(* Logix 5000 project; controller FV vendor 1 type 14 code 217 rev 31.11; software revision 31.00; part 62 of 63 *)
(* tags used below, declared in another part *)
   CWD : CHECKWORD_FLAGS;
   YP_AV1 : PlantItem;   // AV1
   YP_AV2 : PlantItem;   // AV2
   YP_AV3 : PlantItem;   // AV3
   YP_AV4 : PlantItem;   // AV4
   YP_AV5 : PlantItem;   // AV5
   YP_AV6 : PlantItem;   // AV6
   YP_AV7 : PlantItem;   // AV7
   YP_AV8 : PlantItem;   // AV8
   YP_B103 : INT[15];   // Original N File From SLC, No Description Available
   YP_B3 : INT[7];   // BINARY
   YP_B30 : INT[37];   // Original N File From SLC, No Description Available
   YP_B92 : INT[105];   // Original N File From SLC, No Description Available
   YP_BLUNG_OV : PlantItem;   // BLUNG_OV
   YP_C5 : COUNTER[15];
   YP_COMMS_FROM_MVFVCIP : MESSAGE;
   YP_CONV_STOP : PlantItem;   // CONV_STOP
   YP_INP1 : PlantItem;   // INP1
   YP_INP10 : PlantItem;   // INP10
   YP_INP11 : PlantItem;   // INP11
   YP_INP2 : PlantItem;   // INP2
   YP_INP3 : PlantItem;   // INP3
   YP_INP4 : PlantItem;   // INP4
   YP_INP5 : PlantItem;   // INP5
   YP_INP6 : PlantItem;   // INP6
   YP_INP7 : PlantItem;   // INP7
   YP_INP8 : PlantItem;   // INP8
   YP_INP9 : PlantItem;   // INP9
   YP_N14 : INT[135];   // Original N File From SLC, No Description Available
   YP_N40 : INT[9];   // Original N File From SLC, No Description Available
   YP_N55 : INT[244];   // Original N File From SLC, No Description Available
   YP_OUT1 : PlantItem;   // OUT1
   YP_OUT2 : PlantItem;   // OUT2
   YP_OUT3 : PlantItem;   // OUT3
   YP_OUT4 : PlantItem;   // OUT4
   YP_OUT5 : PlantItem;   // OUT5
   YP_OUT6 : PlantItem;   // OUT6
   YP_OUT7 : PlantItem;   // OUT7
   YP_PILZ_OK : PlantItem;   // PILZ_OK
   YP_PRESS_CL : PlantItem;   // PRESS_CL
   YP_PRESS_OP : PlantItem;   // PRESS_OP
   YP_T21 : TIMER[30];
   YP_T4 : TIMER[16];   // TIMER
   YP_WD : PlantItem;   // WD
   YP_WD_RawOutput : ALIAS FOR RIO_Rack_3:3:O.Data.14;   // YP_WD
   YST_BL_PMP_ON : BOOL;   // Blunger Pump
(* YP_Common, continued *)

ROUTINE YP_Digital_Outputs   (* ladder *)
   0: [NEQ(YP_WD.DriveBits,0) OTE(YP_WD.CW.[CWD.AUTODRV]) ,XIC(S:FS) OTU(YP_WD.CW.[CWD.MANUAL]) ,[XIC(YP_WD.CW.[CWD.AUTODRV]) XIO(YP_WD.CW.[CWD.MANUAL]) ,XIC(YP_WD.CW.[CWD.MANDRV]) XIC(YP_WD.CW.[CWD.MANUAL]) ] OTE(YP_WD.CW.[CWD.OUTPUT]) ,XIC(YP_WD.CW.[CWD.OUTPUT]) OTE(YP_WD_RawOutput) ];
END_ROUTINE

ROUTINE YP_INPUTS_10   (* ladder *)
   0: XIC(YP_AV1.CW.[CWD.OPENFB])OTE(YP_B3[0].0);
   1: XIC(YP_AV2.CW.[CWD.OPENFB])OTE(YP_B3[0].2);
   2: XIC(YP_AV3.CW.[CWD.OPENFB])OTE(YP_B3[0].4);
   3: XIC(YP_AV4.CW.[CWD.OPENFB])OTE(YP_B3[0].6);
   4: XIC(YP_AV5.CW.[CWD.OPENFB])OTE(YP_B3[0].8);
   5: XIC(YP_AV6.CW.[CWD.OPENFB])OTE(YP_B3[0].10);
   6: XIC(YP_AV7.CW.[CWD.OPENFB])OTE(YP_B3[0].12);
   7: XIC(YP_AV8.CW.[CWD.OPENFB])OTE(YP_B3[0].14);
   8: XIC(YP_PILZ_OK.CW.[CWD.INPUTSTATUS])OTE(YP_B3[1].0);
   9: XIC(YP_BLUNG_OV.CW.[CWD.INPUTSTATUS])OTE(YP_B3[1].1);
   10: XIO(YP_INP1.CW.[CWD.INPUTSTATUS])OTE(YP_B3[1].2);
   11: XIC(YP_INP2.CW.[CWD.INPUTSTATUS])OTE(YP_B3[1].3);
   12: XIC(YP_INP3.CW.[CWD.INPUTSTATUS])OTE(YP_B3[1].4);
   13: XIC(YP_PRESS_CL.CW.[CWD.INPUTSTATUS])OTE(YP_B3[1].5);
   14: XIC(YP_PRESS_OP.CW.[CWD.INPUTSTATUS])OTE(YP_B3[1].6);
   15: XIC(YP_CONV_STOP.CW.[CWD.INPUTSTATUS])OTE(YP_B3[1].7);
   16: XIC(YP_INP4.CW.[CWD.INPUTSTATUS])OTE(YP_B3[1].8);
   17: XIC(YP_INP5.CW.[CWD.INPUTSTATUS])OTE(YP_B3[1].9);
   18: XIC(YP_INP6.CW.[CWD.INPUTSTATUS])OTE(YP_B3[1].10);
   19: XIC(YP_INP7.CW.[CWD.INPUTSTATUS])OTE(YP_B3[1].11);
   20: XIC(YP_INP8.CW.[CWD.INPUTSTATUS])OTE(YP_B3[1].12);
   21: XIC(YP_INP9.CW.[CWD.INPUTSTATUS])OTE(YP_B3[1].13);
   22: XIC(YP_INP10.CW.[CWD.INPUTSTATUS])OTE(YP_B3[1].14);
   23: XIC(YP_INP11.CW.[CWD.INPUTSTATUS])OTE(YP_B3[1].15);
END_ROUTINE

ROUTINE YP_LAD15_15   (* ladder *)
   0: XIO(YP_T4[3].DN)TON(YP_T4[3],?,?);
   1: XIO(YP_N40[0].0)XIO(YP_N40[0].1)XIO(YP_N40[0].2)XIO(YP_N40[0].3)XIO(YP_N40[0].4)XIO(YP_N40[0].5)XIO(YP_N40[0].6)XIO(YP_N40[0].7)XIO(YP_N40[0].8)[OTL(YP_N40[0].0) ,OTU(YP_N40[0].1) ,OTU(YP_N40[0].2) ,OTU(YP_N40[0].3) ,OTU(YP_N40[0].4) ,OTU(YP_N40[0].5) ,OTU(YP_N40[0].6) ,OTU(YP_N40[0].7) ,OTU(YP_N40[0].8) ];
   2: XIC(YP_N40[0].8)XIC(YP_B3[1].7)[OTU(YP_N40[0].8) ,OTL(YP_N40[0].0) ];
   3: XIC(YP_N40[0].0)XIC(YP_B3[1].0)XIC(YP_B3[1].5)EQU(YP_N55[0],0)[OTU(YP_N40[0].0) ,OTL(YP_N40[0].1) ];
   4: XIC(YP_N40[0].1)XIC(YP_B3[1].1)[OTU(YP_N40[0].1) ,OTL(YP_N40[0].2) ];
   5: XIC(YP_N40[0].2)TON(YP_T21[0],?,?);
   6: XIC(YP_N40[0].2)XIC(YP_T21[0].DN)[OTU(YP_N40[0].2) ,OTL(YP_N40[0].3) ];
   7: MOV(YP_N55[20],YP_C5[0].PRE);
   8: XIC(YP_N40[0].3)XIC(YP_T4[3].DN)CTU(YP_C5[0],?,?);
   9: [XIC(YP_C5[0].DN) ,XIC(YP_C5[1].DN) ][XIC(YP_N40[0].3) ,XIC(YP_B103[4].0) ][OTU(YP_N40[0].3) ,OTL(YP_N40[0].4) ];
   10: MOV(YP_N55[21],YP_C5[1].PRE);
   11: XIC(YP_T4[3].DN)[XIC(YP_N40[0].3) ,XIC(YP_N40[0].4) ]CTU(YP_C5[1],?,?);
   12: XIC(YP_N40[0].4)[XIC(YP_C5[1].DN) ,XIC(YP_B3[1].4) ,XIC(YP_B103[4].0) ][OTU(YP_N40[0].4) ,OTL(YP_N40[0].5) ];
   13: MOV(YP_N55[22],YP_C5[2].PRE);
   14: XIC(YP_T4[3].DN)XIC(YP_N40[0].5)CTU(YP_C5[2],?,?);
   15: XIC(YP_N40[0].5)XIC(YP_C5[2].DN)[OTU(YP_N40[0].5) ,OTL(YP_N40[0].6) ];
   16: XIC(YP_N40[0].6)XIC(YP_B3[1].6)[OTU(YP_N40[0].6) ,OTL(YP_N40[0].7) ];
   17: XIC(YP_N40[0].7)XIC(YP_B3[1].2)[OTU(YP_N40[0].7) ,OTL(YP_N40[0].8) ];
   18: XIC(YP_N40[0].0)[RES(YP_C5[0]) ,RES(YP_C5[1]) ,RES(YP_C5[2]) ];
   19: XIC(YP_N40[0].5)OTU(YP_B103[4].0);
END_ROUTINE

ROUTINE YP_LAD16_16   (* ladder *)
   0: [XIO(YP_N40[1].0) XIO(YP_N40[1].1) XIO(YP_N40[1].2) XIO(YP_N40[1].3) XIO(YP_N40[1].4) XIO(YP_N40[1].5) ,XIC(YP_N40[1].0) NEQ(YP_N55[0],1) ]OTL(YP_N40[1].0);
   1: XIC(YP_N40[1].5)XIC(YP_B3[1].2)[OTU(YP_N40[1].5) ,OTL(YP_N40[1].0) ];
   2: XIC(YP_N40[1].0)XIC(YP_B3[1].0)XIC(YP_B3[1].5)EQU(YP_N55[0],1)[OTU(YP_N40[1].0) ,OTL(YP_N40[1].1) ];
   3: XIC(YP_N40[1].1)XIC(YP_B3[1].1)[OTU(YP_N40[1].1) ,OTL(YP_N40[1].2) ];
   4: XIC(YP_N40[1].2)EQU(YP_N55[10],3)EQU(YP_N55[11],36)XIC(YP_N14[4].1)OTL(YP_B103[2].2);
   5: XIC(YP_N40[1].2)EQU(YP_N55[14],3)EQU(YP_N55[15],36)XIC(YP_N14[14].1)OTL(YP_B103[2].3);
   6: XIC(YP_N40[1].2)[XIC(YP_B103[2].2) ,XIC(YP_B103[2].3) ][OTU(YP_N40[1].2) ,OTL(YP_N40[1].3) ];
   7: XIC(YP_T4[3].DN)XIC(YP_N40[1].3)CTU(YP_C5[10],?,?);
   8: [XIC(YP_N40[1].0) ,GEQ(YP_C5[10].ACC,YP_N55[13]) ]RES(YP_C5[10]);
   9: XIC(YP_N40[1].3)LES(YP_C5[10].ACC,YP_N55[12])OTE(YP_B103[2].0);
   10: XIC(YP_N40[1].3)GEQ(YP_C5[10].ACC,YP_N55[12])OTE(YP_B103[2].1);
   11: XIC(YP_N40[1].3)[XIC(YP_B103[2].2) XIC(YP_N14[4].3) ,XIC(YP_B103[2].3) XIC(YP_N14[14].3) ][OTU(YP_N40[1].3) ,OTL(YP_N40[1].4) ,OTU(YP_B103[2].2) ,OTU(YP_B103[2].3) ];
   12: XIC(YP_N40[1].4)XIC(YP_B3[1].6)XIO(YP_N14[4].0)[OTU(YP_N40[1].4) ,OTL(YP_N40[1].5) ];
END_ROUTINE

ROUTINE YP_LAD20_20   (* ladder *)
   0: XIO(YP_T4[0].DN)TON(YP_T4[0],?,?);
   1: LES(YP_T4[0].ACC,2000)AFI()MSG(YP_COMMS_FROM_MVFVCIP);
   2: XIC(YP_N14[0].0)OTE(YP_N14[100].0);
   3: XIC(YP_N14[0].0)TON(YP_T4[1],?,?);
   4: XIO(YP_N14[0].0)TON(YP_T4[2],?,?);
   5: [XIC(YP_T4[1].DN) ,XIC(YP_T4[2].DN) ]OTE(YP_B103[0].0);
   6: MOV(YP_N14[1],YP_N55[10]);
   7: MOV(YP_N14[2],YP_N55[11]);
   8: MOV(YP_N14[11],YP_N55[14]);
   9: MOV(YP_N14[12],YP_N55[15]);
   10: XIC(YP_B3[1].0)[XIC(YP_N40[1].2) ,XIC(YP_N40[1].3) ]XIO(YP_B103[0].0)[OTE(YP_N14[101].0) ,OTE(YP_N14[111].0) ];
   11: XIC(YP_B3[1].0)XIC(YP_N40[1].3)XIO(YP_B103[0].0)[OTE(YP_N14[104].0) ,OTE(YP_N14[114].0) ];
   12: XIC(YP_N40[1].4)[OTE(YP_N14[104].1) ,OTE(YP_N14[114].1) ];
   13: [MOV(0,YP_N14[103]) ,MOV(0,YP_N14[113]) ];
   14: [XIC(YP_B92[0].0) ,XIC(YP_B92[0].1) ][MOV(3000,YP_N14[103]) ,MOV(3000,YP_N14[113]) ];
   15: [XIC(YP_B92[0].2) ,XIC(YP_B92[0].3) ][MOV(3001,YP_N14[103]) ,MOV(3001,YP_N14[113]) ];
   16: [XIC(YP_B92[0].4) ,XIC(YP_B92[0].5) ][MOV(3002,YP_N14[103]) ,MOV(3002,YP_N14[113]) ];
   17: [XIC(YP_B92[0].6) ,XIC(YP_B92[0].7) ][MOV(3003,YP_N14[103]) ,MOV(3003,YP_N14[113]) ];
   18: [XIC(YP_B92[0].8) ,XIC(YP_B92[0].9) ][MOV(3004,YP_N14[103]) ,MOV(3004,YP_N14[113]) ];
   19: [XIC(YP_B92[0].10) ,XIC(YP_B92[0].11) ][MOV(3005,YP_N14[103]) ,MOV(3005,YP_N14[113]) ];
   20: [XIC(YP_B92[0].12) ,XIC(YP_B92[0].13) ][MOV(3006,YP_N14[103]) ,MOV(3006,YP_N14[113]) ];
   21: [XIC(YP_B92[0].14) ,XIC(YP_B92[0].15) ][MOV(3007,YP_N14[103]) ,MOV(3007,YP_N14[113]) ];
   22: XIO(YP_B3[1].0)[MOV(3011,YP_N14[103]) ,MOV(3011,YP_N14[113]) ];
END_ROUTINE

ROUTINE YP_OUTPUTS_11   (* ladder *)
   0: XIC(YP_B30[0].0)XIC(YP_B3[1].6)XIC(YP_B3[1].0)XIO(YP_B3[1].8)XIO(YP_OUT2.CW.[CWD.OUTPUT])OTE(YP_OUT1.DriveBits.0);
   1: XIC(YP_B30[0].1)XIC(YP_B3[1].5)XIC(YP_B3[1].0)XIO(YP_B3[1].8)XIO(YP_OUT1.CW.[CWD.OUTPUT])OTE(YP_OUT2.DriveBits.0);
   2: XIC(YP_B30[0].2)XIC(YP_B3[1].0)XIO(YP_B3[1].9)XIC(YP_B3[1].14)OTE(YP_OUT3.DriveBits.0);
   3: XIC(YP_B30[0].3)OTE(YP_AV1.DriveBits.0);
   4: XIC(YP_B30[0].4)XIC(YP_B3[1].0)OTE(YP_OUT4.DriveBits.0);
   // Enable Blunger (Wilden) Pump
   5: [XIC(YP_B30[0].5) ,XIC(YST_BL_PMP_ON) ]OTE(YP_AV2.DriveBits.0);
   6: XIC(YP_B30[0].6)OTE(YP_AV3.DriveBits.0);
   7: XIC(YP_B30[0].7)OTE(YP_AV4.DriveBits.0);
   8: XIC(YP_B30[0].8)OTE(YP_AV5.DriveBits.0);
   9: XIC(YP_B30[0].9)XIC(YP_B3[1].0)OTE(YP_AV6.DriveBits.0);
   10: XIC(YP_B30[0].10)XIC(YP_B3[1].0)OTE(YP_AV7.DriveBits.0);
   11: XIC(YP_B30[0].11)XIC(YP_B3[1].0)OTE(YP_AV8.DriveBits.0);
   12: XIC(YP_B30[0].12)XIC(YP_B3[1].0)OTE(YP_OUT5.DriveBits.0);
   13: XIC(YP_B30[0].13)XIC(YP_B3[1].0)OTE(YP_OUT6.DriveBits.0);
   14: XIC(YP_B30[0].14)XIC(YP_B3[1].0)OTE(YP_WD.DriveBits.0);
   15: [XIC(YP_OUT1.CW.[CWD.OUTPUT]) ,XIC(YP_OUT2.CW.[CWD.OUTPUT]) ]XIC(YP_B3[1].0)TON(YP_T4[10],?,?);
   16: [XIC(YP_B30[0].15) ,XIC(YP_T4[10].DN) ]XIC(YP_B3[1].0)OTE(YP_OUT7.DriveBits.0);
   17: XIC(YP_N40[0].6)MOV(1,YP_N55[1]);
   18: XIO(YP_N40[0].6)MOV(0,YP_N55[1]);
END_ROUTINE
